// Mitsubishi GX Works2 project: ZhaoQing_OCV__5.13   PLC: Q10UDEH

TYPE ConveyorIO : STRUCT
  xUnloadCCW : BOOL;  (* 下料为反转 *)
  xUnloadAlarm : BOOL;  (* 下料报警 *)
  xUnload : BOOL;  (* 下料请求 *)
  xPutInto : BOOL;  (* 线体直接投入物料 *)
  xNotArriveAlarm : BOOL;  (* 未到达报警 *)
  xNextRun : BOOL;  (* 下段线体运行 *)
  xMotorCW : BOOL;  (* 电机正转 *)
  xMotorCCW : BOOL;  (* 电机反转 *)
  xManual : BOOL;  (* 手动 *)
  xloadCCW : BOOL;  (* 上料为反转 *)
  xLimitAlarrm : BOOL;  (* 限位报警 *)
  xLoad : BOOL;  (* 上料请求 *)
  xForward : BOOL;  (* 正转手动 *)
  xEmpty : BOOL;  (* 线体状态为空 *)
  xCWPresent : BOOL;  (* 正转检测有无传感器 *)
  xCCWPresent : BOOL;  (* 反转检测有无传感器 *)
  xBusy : BOOL;  (* 工作中 *)
  xBackward : BOOL;  (* 反转手动 *)
  xAuto : BOOL;  (* 自动 *)
  xPosLimit : BOOL;  (* 正限位 *)
  xNegLimit : BOOL;  (* 负限位 *)
  xOverWidthAlarm : BOOL;  (* 超宽报警 *)
  xError : BOOL;  (* 报警 *)
  iProductCategoryIn : INT;  (* 产品类型输入 *)
  iProductCategory : INT;  (* 产品类型记录 *)
  iProductCategoryOut : INT;  (* 产品类型输出 *)
  iDeviceID : INT;  (* 设备编号 *)
  tUnloadAlarmDelay : TIME;  (* 下料报警时间设置 *)
  tLoadDelay : TIME;  (* 上料延时设置 *)
  xSizeDeficientDetect : BOOL;  (* 尺寸缺陷检测 *)
  uiTaskIDIn : WORD;  (* 任务ID输入 *)
  uiTaskID : WORD;  (* 任务ID记录 *)
  uiTaskIDOut : WORD;  (* 任务ID输出 *)
  uiDestinationAdrIn : WORD;  (* 目标地址输入 *)
  uiDestinationAdr : WORD;  (* 目标地址记录 *)
  uiDestinationAdrOut : WORD;  (* 目标地址输出 *)
END_STRUCT END_TYPE

TYPE ShuttleCarIO : STRUCT
  xReady : BOOL;  (* 准备就绪 *)
  xForward : BOOL;  (* 正转 *)
  xBackward : BOOL;  (* 反转 *)
  iCurrentPos : INT;  (* 当前位置 *)
  iDestinationPos : INT;  (* 目标位置 *)
  xCW : BOOL;  (* 正转输出 *)
  xCCW : BOOL;  (* 反转输出 *)
  xBrake : BOOL;  (* 刹车 *)
  xHomeSwitch : BOOL;  (* 零位接近开关 *)
  xPosLimit : BOOL;  (* 正限位 *)
  xNegLimit : BOOL;  (* 负限位 *)
  xMDIExe : BOOL;  (* MDI开始 *)
  xMDIDone : BOOL;  (* MDI 完成 *)
  xPassLimit : BOOL;  (* 限位屏蔽 *)
  xPosLimitCatch : BOOL;  (* 正限位捕捉 *)
  xNegLimitCatch : BOOL;  (* 负限位捕捉 *)
  xHomeExe : BOOL;  (* 开始寻零 *)
  xHomeDone : BOOL;  (* 寻零完成 *)
  xHomeBusy : BOOL;  (* 寻零中 *)
  xHomeFailed : BOOL;  (* 寻零失败 *)
  xBusy : BOOL;  (* 工作中 *)
  tArriveDelay : TIME;  (* 到位延时 *)
  xCylinder : BOOL;  (* 气缸控制 *)
  tBrakeDelay : TIME;  (* 抱闸延时 *)
  xPauseRamp : BOOL;  (* 暂停减速斜坡标志位 *)
  xPresentDetect1 : BOOL;  (* 物料有无检测1 *)
  xPresentDetect2 : BOOL;  (* 物料有无检测2 *)
  xOvertimeAlarm : BOOL;  (* 超时报警 *)
  tSetOverTime : TIME;  (* 设置超时时间 *)
  xLooseDetect : BOOL;  (* 松绳检测 *)
  xLooseAlarm : BOOL;  (* 松绳报警 *)
END_STRUCT END_TYPE

TYPE SwitchIO : STRUCT
  xLiftCylinderRetractDetect : BOOL;
  xLiftCylinderExtendDetect : BOOL;
  xLiftCylinderRetract : BOOL;
  xLiftCylinderExtend : BOOL;
  xEntryBarCylinderRetract : BOOL;
  xLiftCylinderExtendInit : BOOL;
  xEntryEnable : BOOL;
  xExitEnable : BOOL;
  xExitBarCylinderRetract : BOOL;
  xSwithEnable : BOOL;
  xLiftCylinderRetractButton : BOOL;
  xLiftCylinderExtendButton : BOOL;
  xEntryBarCylinderRetractButton : BOOL;
  xExitBarCylinderRetractButton : BOOL;
  xPutInto : BOOL;  (* 单体复位 *)
  tSetOvertime : TIME;  (* 设定超时报警时间 *)
  xOvertimeAlarm : BOOL;  (* 超时报警 *)
END_STRUCT END_TYPE

TYPE BarCylinderIO : STRUCT
  xBarCylinderButton : BOOL;  (* 阻挡气缸 *)
  xPresentSwitch : BOOL;  (* 行程开关 *)
  xBarCylinder : BOOL;  (* 阻挡气缸 *)
  xLoad : BOOL;  (* 上料 *)
  xEmpty : BOOL;  (* 为空指示 *)
  xNextRun : BOOL;  (* 下位设备开始运行 *)
  xUnload : BOOL;  (* 下料 *)
  xTransportMotorCWButton : BOOL;  (* 输送电机正转按钮 *)
  xTransportMotorCW : BOOL;  (* 输送电机正转 *)
  xTransportMotorCCWButton : BOOL;  (* 输送电机反转按钮 *)
  xTransportMotorCCW : BOOL;  (* 输送电机反转 *)
  iProductCategory : INT;  (* 产品种类 *)
  tLoadDelay : TIME;  (* 上料延时 *)
END_STRUCT END_TYPE

// global labels: Global1
VAR_GLOBAL
  g_xAuto AT M11 : BOOL;
  g_xManual : BOOL;
  g_xEStop AT X0BC : BOOL;
  g_xReset AT X0BE : BOOL;
  g_xStackLampRed AT Y2C1 : BOOL;
  g_xStackLampAmber AT Y2C3 : BOOL;
  g_xStackLampGreen AT Y2C2 : BOOL;
  g_xBuzzer AT Y2C4 : BOOL;
  g_xStop AT M2 : BOOL;
  g_xLocalAutoStart AT M1 : BOOL;
  g_xRemoteAutoStart AT M0 : BOOL;
  g_xRemoteAuto AT M10 : BOOL;
  g_iState AT D40 : INT;
  g_iLocalAutoStep : BOOL;
  g_xAlarm : BOOL;
  g_xPause AT M3 : BOOL;  (* 暂停 *)
  g_iDeviceIDSelect AT D0 : INT;
  g_xImport1Force AT M165 : BOOL;
  g_xImport2Force AT M166 : BOOL;
  g_xImport3Force AT M167 : BOOL;
  g_xResetSingle AT M4 : BOOL;  (* 单线体复位 *)
  g_xInsertTask AT M5 : BOOL;  (* 插入任务 *)
  g_iInsertTask AT D2 : INT;  (* 插入任务号 *)
  g_iConveyorStatus AT D4 : INT;
  g_xChenPinComFailed AT M168 : BOOL;
END_VAR

// task Task_01 (event TRUE, interval 0, priority 31): POU, Start, tcp

FUNCTION_BLOCK Conveyor
VAR
  m_xPresentDelay : BOOL;  (* 有无判断延时 *)
  m_xLoadDelayOut : BOOL;  (* 上料延时输出 *)
  m_xInitial : BOOL;  (* 初始化 *)
  m_tUnloadTimer : TIME;  (* 下料计时器 *)
  m_tPresentDelayCurrentTime : TIME;
  m_tonUnloadAlam : TON;  (* 下料报警定时器 *)
  m_tonPresentDelay : TON;  (* 物料有无判断延时，防止误动作 *)
  m_tonNotArriveAlarm : TON;  (* 未到达报警计时 *)
  m_tonLoadDelay : TON;  (* 上料延时 *)
  m_tNotArriveCurrentTime : TIME;  (* 未到达报警计时当前时间 *)
  m_tLoadTimer : TIME;  (* 上料计时器 *)
  iStep : INT;  (* 上料步骤 *)
  m_wStateWord : INT;
END_VAR
VAR_IN_OUT
  ConveyorMotor : ConveyorIO;  (* 输送线输入输出 *)
END_VAR
(*////////////////////////////////////////////////////////////////////////////////////////////////////////////
//传输线控制FB块，可控制单方向线体，双向旋转线体，支持双向上下料            
//线体初始化后为空的情况下输入xLoad信号即可进行上料动作，使用xLoadCCW信号可反方向上料
//增加了产品信息和产品种类的储存，当传输线为空和上料进行标志位为零的情况下清除产品信息和产品种类
//使用方式是在置位xLoad信号后，把产品信息和产品种类传入，等下料后自动清零
//线体不为空的情况下使用xUnload信号可进行下料动作，物料有无传感器的下降沿后出发计时器，延时断开传输线旋转
//单方向传输线体把xLoadCCW、xUnloadCCW设置为零，双向线体上料方向和下料反向的,方向固定的 把xUnloadCCW设置为1
//双方向线体双向都能上下料的要根据上料的方向来设置xLoadCCW,xUnloadCCW
//增加工作中信号xBusy当电机正转 显示为工作中
//增加上下料超时报警，xLoadAlarm，xUnloadAlarm，设定时间在LOAD_UNLOAD_TIME常量上，现在设置的为30秒
//增加xPutInto信号，用于直接投入的物料，检测开关感应到后，直接进入下料流程，上升沿有效
//离开延时改为变量 iLeaveDelay 默认为0 离开检测开关离输送线尾端比较远的线体需要根据情况设定100ms为单位
//增加初始化标志位，增加进入延时时间，初始化为进入延时时间为0 ，离开延时时间为2S，通过外围接口可以更改
//修改信息  修改后请增加版本
//12-17进行了优化，增加了未到达报警，当物料未传送到下一设备，就报未到达报警，使用xNextRun标志位制作，没有正常到达
//第0步，不能跳转到第一步把标志位复位，即出现中断情况，2秒后报警
//修改信息  修改后请增加版本
上料延时增加为50ms防止干扰信号
nextrun信号在 第三步也要复位
增加限位报警
增加超宽报警
增加产品型号输出在下料的时候把产品型号输送给下一段线体
增加线体单独复位
增加任务插入功能配合全局变量
增加暂停功能
增加线体状态字显示  0 空闲 1：有料  2 工作中  3  超限报警 4 超宽报警  5 未到达报警  6 下料超时报警
空料判断放在自动前，进行有无报警判断，然后跳转
//YAO      V1.0
///////////////////////////////////////////////////////////////////////////////////////////////////////////
(*********************************************************)
(*//初始化，
//上料延时位0S，下料报警延时为30S
//下料延时设一个比较大的时间，主要依靠xunload标志位来停止输送线，特殊情况可以用延时来停止物流线下料
//设置时间大的时候计时器会失效*)
IF NOT m_xInitial THEN
	ConveyorMotor.tLoadDelay:=T#100ms;
	ConveyorMotor.tUnloadAlarmDelay:=T#30s;
	ConveyorMotor.xPosLimit:=1;
	ConveyorMotor.xNegLimit:=1;
	ConveyorMotor.xSizeDeficientDetect:=0;
	m_xInitial:=1;
END_IF;
(*//自动
//复位信号把步号置0，但xLoad与xUnload没有复位，调用程序需要注意复位后把这两个信号置零，以免发生误动作
//物料有无判断增加延时，防止开自动瞬间误动作发生*)
m_tonPresentDelay(IN:= ConveyorMotor.xCWPresent OR ConveyorMotor.xCCWPresent,
                  PT:=T#100ms,
				  Q:= m_xPresentDelay,
				  ET:= m_tPresentDelayCurrentTime);
CASE iStep OF
	0:(*//初始化*)
	ConveyorMotor.xMotorCW:=0;
	ConveyorMotor.xMotorCCW:=0;
	ConveyorMotor.iProductCategoryOut:=0;
	ConveyorMotor.uiTaskIDOut:=0;
	ConveyorMotor.uiDestinationAdOut:=0;
(*	//判断物料有无传感器*)	
		IF m_xPresentDelay THEN			
			ConveyorMotor.xEmpty:=0;
			IF g_xAuto AND NOT ConveyorMotor.xError THEN(*//自动情况下进行跳转*)(*无超限报警*)
				iStep:=3;
			END_IF;
		ELSE
			ConveyorMotor.xEmpty:=1;
			IF g_xAuto AND NOT ConveyorMotor.xError THEN(*//自动情况下进行跳转*)(*无超限报警*)
				iStep:=1;	
			END_IF;		
	END_IF;	
	1: (*//上料*)
	ConveyorMotor.xNextRun:=0;
	IF ConveyorMotor.xLoad    THEN (*//上料开始*)
		ConveyorMotor.iProductCategory:=0;	(*//上料开始清除产品信息*)
		ConveyorMotor.uiTaskID:=0;
		ConveyorMotor.uiDestinationAdr:=0;		
		iStep:=2;		
	END_IF;
	2: (*//上料完成*)
	ConveyorMotor.iProductCategory:=ConveyorMotor.iProductCategoryIn;(* //产品信息传入*)		
	ConveyorMotor.uiTaskID:=ConveyorMotor.uiTaskIDIn;
	ConveyorMotor.uiDestinationAdr:=ConveyorMotor.uiDestinationAdrIn;
	IF ConveyorMotor.xloadCCW THEN
		ConveyorMotor.xMotorCCW:=1; 
		ConveyorMotor.xMotorCW:=0;
	ELSE
	    ConveyorMotor.xMotorCW:=1;  
		ConveyorMotor.xMotorCCW:=0;
	END_IF;
		m_tonLoadDelay(IN:= (ConveyorMotor.xCWPresent AND NOT ConveyorMotor.xloadCCW) 
		                                        OR (ConveyorMotor.xCCWPresent AND ConveyorMotor.xloadCCW) ,
		                               PT:= ConveyorMotor.tLoadDelay ,
		                               Q:= m_xLoadDelayOut ,
		                               ET:= m_tLoadTimer );
	    IF (m_xLoadDelayOut AND NOT ConveyorMotor.xSizeDeficientDetect)   (*无尺寸检测时  只检测一个开关*)
	    	OR (m_xLoadDelayOut AND ConveyorMotor.xSizeDeficientDetect(*有尺寸检测时  要检测两个开关*)
	    	                                          AND ConveyorMotor.xCCWPresent 
	    	                                          AND ConveyorMotor.xCWPresent)      THEN 	 
		    iStep:=3;
			    ELSIF (m_xLoadDelayOut 
		                       AND ConveyorMotor.xSizeDeficientDetect(*尺寸不足报警*)
	    	                  AND (NOT ConveyorMotor.xCCWPresent OR NOT ConveyorMotor.xCWPresent))  
	    THEN
	    	    ConveyorMotor.xOverWidthAlarm:=1;
	    	   iStep:=0;               
	    END_IF;

	3:(*//下料请求*)	
	ConveyorMotor.xMotorCW:=0;
	ConveyorMotor.xMotorCCW:=0;
	ConveyorMotor.xEmpty:=0;
	IF ConveyorMotor.xUnload AND NOT ConveyorMotor.xOverWidthAlarm  THEN (*无超宽报警可以下料*)
		iStep:=4;
	END_IF;
	4:(*	//下料完成*)
	IF ConveyorMotor.xUnloadCCW THEN   
		ConveyorMotor.xMotorCCW:=1;  
		ConveyorMotor.xMotorCW:=0;
		ELSE
	    ConveyorMotor.xMotorCW:=1;  
		ConveyorMotor.xMotorCCW:=0;
	END_IF;
	ConveyorMotor.xNextRun:=1; (*下一段线体旋转*)
	ConveyorMotor.iProductCategoryOut:=ConveyorMotor.iProductCategory;(*产品型号输出给下一段线体*)
	ConveyorMotor.uiDestinationAdrOut:=ConveyorMotor.uiDestinationAdr;
	ConveyorMotor.uiTaskIDOut:=
	IF NOT ConveyorMotor.xUnload THEN 
		istep:=0;
	END_IF;
END_CASE;
(*投入上料，搬出下料，也可用来初始化*)
IF LDP(TRUE,ConveyorMotor.xPutInto) THEN
	iStep:=0;
END_IF;
(*//当前任务显示*)
IF LDP(TRUE,ConveyorMotor.iDeviceID=g_iDeviceIDSelect) THEN
	g_iInsertTask:=ConveyorMotor.iProductCategory;
END_IF;
	(*//插入任务*)
IF g_xInsertTask AND ConveyorMotor.iDeviceID=g_iDeviceIDSelect THEN
	ConveyorMotor.iProductCategory:=g_iInsertTask;
END_IF;
(*//单线体复位，当设备号与本线体一致的时候执行复位*)
IF (g_xResetSingle AND ConveyorMotor.iDeviceID=g_iDeviceIDSelect)THEN (* //非正常情况下切断xNextRun不会复位，通过这个标志位会出发报警*)(*增加单体复位*)
	iStep:=0;
	ConveyorMotor.xNextRun:=0; 
	ConveyorMotor.xLimitAlarrm:=0;
	ConveyorMotor.xOverWidthAlarm:=0;
END_IF;
(*//手动*)
IF g_xManual THEN
(*	iStep:=0; *)(*//手动后上下料程序步骤清零*)
	(*//正转*)
	IF ConveyorMotor.xForward 
		AND ConveyorMotor.xBackward=0 
		AND ConveyorMotor.xMotorCCW=0 
		AND g_xEStop THEN
		ConveyorMotor.xMotorCW:=1;
		ConveyorMotor.xMotorCCW:=0;
		ELSE
		ConveyorMotor.xMotorCW:=0;
	END_IF;
	(*//反转*)
	IF ConveyorMotor.xBackward 
		AND ConveyorMotor.xForward=0 
		AND ConveyorMotor.xMotorCW=0 
		AND g_xEStop THEN
		ConveyorMotor.xMotorCCW:=1;
		conveyormotor.xMotorCW:=0;
		ELSE
		ConveyorMotor.xMotorCCW:=0;
	END_IF;
END_IF;
(*暂停*)
IF g_xPause THEN
	ConveyorMotor.xMotorCCW:=0;
	ConveyorMotor.xMotorCW:=0;
END_IF;
(*工作中信号输出*)
ConveyorMotor.xBusy:=ConveyorMotor.xMotorCCW OR ConveyorMotor.xMotorCW;
(*//未到达报警*)
m_tonNotArriveAlarm(IN:= iStep=0 AND ConveyorMotor.xNextRun  ,PT:= T#2s,Q:= ConveyorMotor.xNotArriveAlarm ,ET:= m_tNotArriveCurrentTime );
(*//下料超时报警*)
m_tonUnloadAlam(IN:= iStep=4,PT:=ConveyorMotor.tUnloadAlarmDelay,Q:= ConveyorMotor.xUnloadAlarm,ET:=m_tUnloadTimer );
(*//限位报警,进料检测开关失效*)
IF ( ((ConveyorMotor.xloadCCW AND NOT ConveyorMotor.xNegLimit)            (*反转上料，碰到负限位*)
	OR  ( NOT ConveyorMotor.xloadCCW AND NOT ConveyorMotor.xPosLimit)) (*正转上料，碰到正限位*)
    AND iStep=2) (*上料过程*)
    OR
   ( iStep=4 (*下料过程*)
	AND( (ConveyorMotor.xUnloadCCW AND NOT ConveyorMotor.xPosLimit)  
	OR (NOT ConveyorMotor.xUnloadCCW AND NOT ConveyorMotor.xNegLimit)))    
    THEN
    ConveyorMotor.xLimitAlarrm:=1;
    iStep:=0;
END_IF;
(*//超宽报警*)
IF iStep=3 AND (NOT ConveyorMotor.xNegLimit OR NOT ConveyorMotor.xPosLimit) THEN
	ConveyorMotor.xOverWidthAlarm:=1;
END_IF;
(*//总报警*)
ConveyorMotor.xError:=ConveyorMotor.xLimitAlarrm
                                              OR ConveyorMotor.xNotArriveAlarm
                                              OR ConveyorMotor.xUnloadAlarm                                             
                                              OR ConveyorMotor.xOverWidthAlarm;

(*//状态输出*)(*状态显示，容易造成指针容量不足*)
IF ConveyorMotor.xEmpty AND NOT ConveyorMotor.xBusy THEN
	m_wStateWord:=0;
END_IF;
IF ConveyorMotor.xEmpty=0 THEN
		m_wStateWord:=1;
END_IF;
IF ConveyorMotor.xBusy THEN
		m_wStateWord:=2;
END_IF;
IF ConveyorMotor.xLimitAlarrm THEN
		m_wStateWord:=3;
END_IF;
IF ConveyorMotor.xOverWidthAlarm THEN
		m_wStateWord:=4;
END_IF;
(*IF ConveyorMotor.xNotArriveAlarm THEN	
		m_wStateWord:=5;
END_IF;*)
IF ConveyorMotor.xUnloadAlarm THEN
		m_wStateWord:=6;	
END_IF;
(*选择本线体后，将状态赋值给全局变量进行显示*)
IF ConveyorMotor.iDeviceID=g_iDeviceIDSelect THEN
	g_iConveyorStatus:=m_wStateWord;
END_IF;
END_FUNCTION_BLOCK

PROGRAM POU
VAR
  Cylinder12309 : ShuttleCar;
  CylinderIO12309 : ShuttleCarIO;
  ConveyorIO12114 : ConveyorIO;
  Conveyor12114 : Conveyor;
  Conveyor12115 : Conveyor;
  ConveyorIO12115 : ConveyorIO;
  Switch12312 : Switch;
  SwitchIO12312 : SwitchIO;
  Conveyor12123 : Conveyor;
  ConveyorIO12123 : ConveyorIO;
  Conveyor12124 : Conveyor;
  ConveyorIO12124 : ConveyorIO;
  Conveyor12125 : Conveyor;
  ConveyorIO12125 : ConveyorIO;
  Switch12203 : Switch;
  SwitchIO12203 : SwitchIO;
  Conveyor12142 : Conveyor;
  ConveyorIO12142 : ConveyorIO;
  Bar12326 : BarCylinder;
  BarIO12326 : BarCylinderIO;
  Conveyor12116 : Conveyor;
  ConveyorIO12116 : ConveyorIO;
  Cylinder12308 : ShuttleCar;
  CylinderIO12308 : ShuttleCarIO;
  Conveyor12111 : Conveyor;
  ConveyorIO12111 : ConveyorIO;
  Conveyor12112 : Conveyor;
  ConveyorIO12112 : ConveyorIO;
  Switch12311 : Switch;
  SwitchIO12311 : SwitchIO;
  Conveyor12113 : Conveyor;
  ConveyorIO12113 : ConveyorIO;
  Conveyor12120 : Conveyor;
  ConveyorIO12120 : ConveyorIO;
  Conveyor12121 : Conveyor;
  ConveyorIO12121 : ConveyorIO;
  Conveyor12122 : Conveyor;
  ConveyorIO12122 : ConveyorIO;
  Cylinder12307 : ShuttleCar;
  CylinderIO12307 : ShuttleCarIO;
  Conveyor12108 : Conveyor;
  ConveyorIO12108 : ConveyorIO;
  Conveyor12109 : Conveyor;
  ConveyorIO12109 : ConveyorIO;
  Switch12310 : Switch;
  SwitchIO12310 : SwitchIO;
  Conveyor12110 : Conveyor;
  ConveyorIO12110 : ConveyorIO;
  Conveyor12117 : Conveyor;
  ConveyorIO12117 : ConveyorIO;
  Conveyor12118 : Conveyor;
  ConveyorIO12118 : ConveyorIO;
  Conveyor12119 : Conveyor;
  ConveyorIO12119 : ConveyorIO;
  Conveyor12203 : Conveyor;
  ConveyorIO12203 : ConveyorIO;
  Conveyor12143 : Conveyor;
  ConveyorIO12143 : ConveyorIO;
  Switch12330 : Switch;
  ConveyorIO12144 : ConveyorIO;
  ConveyorIO12333 : ConveyorIO;  (* OCV2顶升移载进入线体 *)
  ConveyorIO12152 : ConveyorIO;  (* OCV2顶升移载离开线体 *)
  SwitchIO12333 : SwitchIO;  (* OCV2顶升移载 *)
  m_xTS1ExportPermit : BOOL;  (* OCV2顶升移载 *)
  m_xConveyor12114Export : BOOL;  (* 12114线体输出 *)
  ConveyorIO12146 : ConveyorIO;
  m_xTS2ExportPermit : BOOL;
  m_xMotorFlag : BOOL;
  m_xTS3ExportPermit : BOOL;
  SwitchIO12330 : SwitchIO;
  Switch12333 : Switch;  (* OCV2顶升移载 *)
  SwitchIO12321 : SwitchIO;
  Switch12321 : Switch;  (* OCV2顶升移载 *)
  Conveyor12141 : Conveyor;
  ConveyorIO12141 : ConveyorIO;
  Conveyor12140 : Conveyor;
  ConveyorIO12140 : ConveyorIO;
  m_iSwitch12321Select : INT;
  Conveyor12138 : Conveyor;
  ConveyorIO12138 : ConveyorIO;
  Conveyor12139 : Conveyor;
  ConveyorIO12139 : ConveyorIO;
  Conveyor12136 : Conveyor;
  ConveyorIO12136 : ConveyorIO;
  Conveyor12137 : Conveyor;
  ConveyorIO12137 : ConveyorIO;
  Switch12317 : Switch;
  SwitchIO12317 : SwitchIO;
  ConveyorIO12135 : ConveyorIO;
  ConveyorIO12134 : ConveyorIO;
  m_iSwitch12317Select : INT;
  Conveyor12132 : Conveyor;
  ConveyorIO12132 : ConveyorIO;
  Conveyor12133 : Conveyor;
  ConveyorIO12133 : ConveyorIO;
  Conveyor12131 : Conveyor;
  ConveyorIO12131 : ConveyorIO;
  Conveyor12130 : Conveyor;
  ConveyorIO12130 : ConveyorIO;
  Switch12314 : Switch;
  SwitchIO12314 : SwitchIO;
  Conveyor12129 : Conveyor;
  ConveyorIO12129 : ConveyorIO;
  Conveyor12128 : Conveyor;
  ConveyorIO12128 : ConveyorIO;
  m_iSwitch12314Select : INT;
  Conveyor12126 : Conveyor;
  ConveyorIO12126 : ConveyorIO;
  Conveyor12127 : Conveyor;
  ConveyorIO12127 : ConveyorIO;
  Cylinder12320 : ShuttleCar;
  CylinderIO12320 : ShuttleCarIO;
  Cylinder12316 : ShuttleCar;
  CylinderIO12316 : ShuttleCarIO;
  Cylinder12313 : ShuttleCar;
  CylinderIO12313 : ShuttleCarIO;
  Conveyor12147 : Conveyor;
  ConveyorIO12147 : ConveyorIO;
  Conveyor12148 : Conveyor;
  ConveyorIO12148 : ConveyorIO;
  Lifter8 : ShuttleCar;
  Lifter8IO : ShuttleCarIO;
  Lifter8Speed : ShuttleCarVelocityFB;
  Conveyor8 : Conveyor;
  Conveyor8IO : ConveyorIO;
  Lifter9 : ShuttleCar;
  Lifter9IO : ShuttleCarIO;
  Lifter9Speed : ShuttleCarVelocityFB;
  Conveyor9 : Conveyor;
  Conveyor9IO : ConveyorIO;
  Conveyor12156 : Conveyor;
  ConveyorIO12156 : ConveyorIO;
  Conveyor12155 : Conveyor;
  ConveyorIO12155 : ConveyorIO;
  m_tonSwitch1NOSeleteDelay : TON;
  m_tonSwitch2NOSeleteDelay : TON;
  m_tonSwitch3NOSeleteDelay : TON;
  m_xSwitch12321NoSeleteDelay : BOOL;
  m_xSwitch12317NoSeleteDelay : BOOL;
  m_xSwitch12314NoSeleteDelay : BOOL;
  m_tSwitch12321NOSeleteCurrent : TIME;
  m_tSwitch12317NOSeleteCurrent : TIME;
  m_tSwitch12314NOSeleteCurrent : TIME;
  Switch12312Priority : PriorityFB;
  m_xSwitch12312Task : INT;
  Conveyor12159 : Conveyor;
  ConveyorIO12159 : ConveyorIO;
  Switch12337 : Switch;
  SwitchIO12337 : SwitchIO;
  ConveyorIO12158 : ConveyorIO;
  ConveyorIO12157 : ConveyorIO;
  ConveyorIO12321 : ConveyorIO;
  Switch12311Priority : PriorityFB;
  m_xSwitch12311Task : INT;
  SwitchIO12204 : SwitchIO;
  Switch12204 : Switch;
  ConveyorIO12145 : ConveyorIO;
  ConveyorIO12204 : ConveyorIO;
  Conveyor12151 : Conveyor;
  ConveyorIO12151 : ConveyorIO;
  Conveyor12150 : Conveyor;
  ConveyorIO12150 : ConveyorIO;
  Conveyor12149 : Conveyor;
  ConveyorIO12149 : ConveyorIO;
  Switch12328 : Switch;
  SwitchIO12328 : SwitchIO;
  Lifter8Priority : PriorityFB;
  m_iLifter8Task : INT;
  m_xSwitch12321Select : BOOL;
  m_xSwitch12317Select : BOOL;
  Cylinder12301 : ShuttleCar;
  CylinderIO12301 : ShuttleCarIO;
  Cylinder12302 : ShuttleCar;
  CylinderIO12302 : ShuttleCarIO;
  Cylinder12303 : ShuttleCar;
  CylinderIO12303 : ShuttleCarIO;
  Cylinder12304 : ShuttleCar;
  CylinderIO12304 : ShuttleCarIO;
  Conveyor12101 : Conveyor;
  ConveyorIO12101 : ConveyorIO;
  Conveyor12102 : Conveyor;
  ConveyorIO12102 : ConveyorIO;
  Conveyor12103 : Conveyor;
  ConveyorIO12103 : ConveyorIO;
  Conveyor12104 : Conveyor;
  ConveyorIO12104 : ConveyorIO;
  ShuttleCar12401 : ShuttleCar;
  ShuttleCarIO12401 : ShuttleCarIO;
  Conveyor12105 : Conveyor;
  ConveyorIO12105 : ConveyorIO;
  Conveyor12106 : Conveyor;
  ConveyorIO12106 : ConveyorIO;
  Switch12201 : Switch;
  SwitchIO12201 : SwitchIO;
  Switch12202 : Switch;
  SwitchIO12202 : SwitchIO;
  Conveyor12201 : Conveyor;
  ConveyorIO12201 : ConveyorIO;
  Conveyor12202 : Conveyor;
  ConveyorIO12202 : ConveyorIO;
  Conveyor12401 : Conveyor;
  ConveyorIO12401 : ConveyorIO;
  Rotor12501 : ShuttleCar;
  RotorIO12501 : ShuttleCarIO;
  Conveyor12501 : Conveyor;
  ConveyorIO12501 : ConveyorIO;
  Conveyor12154 : Conveyor;
  ConveyorIO12154 : ConveyorIO;
  ShuttleCar12401Position : ARRAY [0..5] OF INT;
  ii : INT;
  ConveyorIO12107 : ConveyorIO;
  m_xSwitch12314Select : BOOL;
  Conveyor12146 : Conveyor;
  Switch12330ConveyorOut : ConveyorIO;
  m_xPickOutDone : BOOL;  (* 分拣完成 *)
  ConveyorIO12160 : ConveyorIO;  (* OCV1工位 *)
  m_xOCV1Done : BOOL;  (* OCV1完成 *)
  Conveyor12160 : Conveyor;
  Conveyor12161 : Conveyor;
  ConveyorIO12161 : ConveyorIO;
  ConveyorIO12162 : ConveyorIO;
  Conveyor12162 : Conveyor;
  TonScan1 : TON;
  TonScan1Time : TIME;
  TonScan2 : TON;
  TonScan2Time : TIME;
  xTonScan1 : BOOL;
  xTonScan2 : BOOL;
END_VAR
IF M1 AND M2 THEN D333:=D333;END_IF;
(*提升机8*)
Lifter8(ShuttleCarInOut:=Lifter8IO);
(*ShuttleCarCurrentPosition(XC2 OR XC4 OR XC3 ,XC2 ,XC3, XC4, Lifter8IO.iCurrentPos);*)
IF XC1 AND XC2 THEN
	Lifter8IO.iCurrentPos:=1;
ELSIF XC2 AND NOT XC1 THEN
	Lifter8IO.iCurrentPos:=2;
ELSIF XC3 THEN
	Lifter8IO.iCurrentPos:=3;
ELSIF XC4 THEN
	Lifter8IO.iCurrentPos:=4;
END_IF;
Lifter8Speed(xEnable:= g_xAuto,
                        xMotorCW:= Lifter8IO.xCW ,
                        xMotorCCW:= Lifter8IO.xCCW,
                        xPosition1Switch:= XC2 OR XC4,
                        xDecelerationSwitch:= XC0 ,
	                    xPosition2Switch:= XC3 ,
	                   xHighSpeed:= Y296 );
Lifter8IO.xReady:=XBA;
Lifter8IO.xLooseDetect:=XC6;;
Lifter8IO.xForward:=M107 OR XC7;
Lifter8IO.xBackward:=M108 OR XC8;
Lifter8IO.xPosLimit:=XBF;
Lifter8IO.xNegLimit:=XC5;
Y294:=Lifter8IO.xCW;
Y295:=Lifter8IO.xCCW;
Y299:=Lifter8IO.xBrake;
Lifter8IO.tArriveDelay:=T#500ms;

Conveyor8(ConveyorMotor:=Conveyor8IO);
Conveyor8IO.xForward:=M109;
Conveyor8IO.xBackward:=M110;
Conveyor8IO.xCWPresent:=XC9;
Conveyor8IO.xCCWPresent:=XCA;
Y29A:=Conveyor8IO.xMotorCW;
Y29B:=Conveyor8IO.xMotorCCW;
Conveyor8IO.xSizeDeficientDetect:=1;
Conveyor8IO.iDeviceID:=8;

(*提升机9*)
Lifter9(ShuttleCarInOut:=Lifter9IO);
ShuttleCarCurrentPosition(XCC OR XCD ,XCC ,XCD,FALSE, Lifter9IO.iCurrentPos);
Lifter9Speed(xEnable:= g_xAuto,
                        xMotorCW:= Lifter9IO.xCW ,
                        xMotorCCW:=Lifter9IO.xCCW,
                        xPosition1Switch:= XCC,
                        xDecelerationSwitch:= XCB,
	                    xPosition2Switch:= XCD ,
	                    xHighSpeed:= Y2A1 );
Lifter9IO.xReady:=XBB;
Lifter9IO.xForward:=M111 OR XD1;
Lifter9IO.xBackward:=M112 OR XD2;
Lifter9IO.xLooseDetect:=XD0;
Lifter9IO.xPosLimit:=XCE;
Lifter9IO.xNegLimit:=XCF;
Y29F:=Lifter9IO.xCW;
Y2A0:=Lifter9IO.xCCW;
Y2A4:=Lifter9IO.xBrake;

Conveyor9(ConveyorMotor:=Conveyor9IO);
Conveyor9IO.xForward:=M113;
Conveyor9IO.xBackward:=M114;
Conveyor9IO.xCWPresent:=XD4;
Conveyor9IO.xCCWPresent:=XD3;
Y2A6:=Conveyor9IO.xMotorCW;
Y2A5:=Conveyor9IO.xMotorCCW;
Conveyor9IO.iDeviceID:=9;
(*H750高温库人工换内衬线体*)
(*高位库2巷道入库*)
Cylinder12301(ShuttleCarInOut:=CylinderIO12301);
ShuttleCarCurrentPosition( X3 OR X4 ,X4 ,X3, FALSE, CylinderIO12301.iCurrentPos );
CylinderIO12301.xForward:=M137;
CylinderIO12301.xBackward:=M138;
CylinderIO12301.xCylinder:=1;
Y201:=CylinderIO12301.xCW;
Y202:=CylinderIO12301.xCCW;
CylinderIO12301.xPresentDetect1:=X02;

Conveyor12101(ConveyorMotor:=ConveyorIO12101);
ConveyorIO12101.xForward:=M139;
ConveyorIO12101.xCWPresent:=X1;
Y203:=ConveyorIO12101.xMotorCW;
M362:= NOT ConveyorIO12101.xEmpty;
M363:=ConveyorIO12101.xError;
ConveyorIO12101.iDeviceID:=12101;

(*高位库2巷道出库*)
Cylinder12302(ShuttleCarInOut:=CylinderIO12302);
ShuttleCarCurrentPosition( X6 OR X7 ,X7,X6, FALSE, CylinderIO12302.iCurrentPos );
CylinderIO12302.xForward:=M140;
CylinderIO12302.xBackward:=M141;
CylinderIO12302.xCylinder:=1;
Y204:=CylinderIO12302.xCW;
Y205:=CylinderIO12302.xCCW;
CylinderIO12302.xPresentDetect1:=X05;

Conveyor12102(ConveyorMotor:=ConveyorIO12102);
ConveyorIO12102.xForward:=M141;
ConveyorIO12102.xCWPresent:=X8;
Y206:=ConveyorIO12102.xMotorCW;
M410:= NOT conveyorIO12102.xEmpty;
M411:= ConveyorIO12102.xError;
ConveyorIO12102.iDeviceID:=12102;

(*高位库1巷道出库*)
Cylinder12303(ShuttleCarInOut:=CylinderIO12303);
ShuttleCarCurrentPosition( X9 OR XA ,XA,X9, FALSE, CylinderIO12303.iCurrentPos );
CylinderIO12303.xForward:=M142;
CylinderIO12303.xBackward:=M143;
CylinderIO12303.xCylinder:=1;
Y207:=CylinderIO12303.xCW;
Y208:=CylinderIO12303.xCCW;
CylinderIO12303.xPresentDetect1:=X0B;

Conveyor12103(ConveyorMotor:=ConveyorIO12103);
ConveyorIO12103.xForward:=M144;
ConveyorIO12103.xCWPresent:=XC;
M412:= NOT conveyorIO12103.xEmpty;
M413:= ConveyorIO12103.xError;
ConveyorIO12103.iDeviceID:=12103;
Y209:=ConveyorIO12103.xMotorCW;

(*高位库1巷道入库*)
Cylinder12304(ShuttleCarInOut:=CylinderIO12304);
ShuttleCarCurrentPosition( XF OR X10 ,X10,XF, FALSE, CylinderIO12304.iCurrentPos );
CylinderIO12304.xForward:=M145;
CylinderIO12304.xBackward:=M146;
CylinderIO12304.xCylinder:=1;
Y21A:=CylinderIO12304.xCW;
Y21B:=CylinderIO12304.xCCW;
CylinderIO12304.xPresentDetect1:=X0E;

Conveyor12104(ConveyorMotor:=ConveyorIO12104);
ConveyorIO12104.xForward:=M144;
ConveyorIO12104.xCWPresent:=XD;
Y21C:=ConveyorIO12104.xMotorCW;
M414:= NOT conveyorIO12104.xEmpty;
M415:= ConveyorIO12104.xError;
ConveyorIO12104.iDeviceID:=12104;

(*高位库RGV*)
(*ShuttleCar12401(ShuttleCarInOut:= ShuttleCarIO12401 );
ShuttleCar12401Position[0]:=1;
ShuttleCar12401Position[1]:=1;
ShuttleCar12401Position[2]:=1;
ShuttleCar12401Position[3]:=1;
ShuttleCar12401Position[4]:=1;
ShuttleCar12401Position[5]:=1;

Y2CA:=ShuttleCarVelocityEncoder( g_xAuto , D190 , ShuttleCar12401Position[ShuttleCarIO12401.iDestinationPos] );
IF LDP(TRUE,g_xAuto) THEN
	ShuttleCarIO12401.iCurrentPos:=0;
END_IF;
FOR ii:=0 TO 5 BY 1 DO
	IF abs(D190-ShuttleCar12401Position[ii])<10 THEN
		ShuttleCarIO12401.iCurrentPos:=ii;
	END_IF;
END_FOR;

ShuttleCarIO12401.xReady:=XBD;
ShuttleCarIO12401.xForward:=M147 OR XD5;
ShuttleCarIO12401.xBackward:=M148 OR XD6;
ShuttleCarIO12401.xPosLimit:=XDA;
ShuttleCarIO12401.xNegLimit:=XDB;
Y2C8:=ShuttleCarIO12401.xCW;
Y2C9:=ShuttleCarIO12401.xCCW;
Y2BD:=ShuttleCarIO12401.xBrake;

Conveyor12105(ConveyorMotor:=ConveyorIO12105);
ConveyorIO12105.xForward:=M149;
ConveyorIO12105.xCWPresent:=X11;
Y21D:=ConveyorIO12105.xMotorCW;
M416:= NOT conveyorIO12105.xEmpty;
M417:= ConveyorIO12105.xError;
ConveyorIO12105.iDeviceID:=12105;

Conveyor12106(ConveyorMotor:=ConveyorIO12106);
ConveyorIO12106.xForward:=M150;
ConveyorIO12106.xCWPresent:=X12;
Y21E:=ConveyorIO12106.xMotorCW;
M418:= NOT conveyorIO12106.xEmpty;
M419:= ConveyorIO12106.xError;
ConveyorIO12106.iDeviceID:=12106;

Switch12202(ConveyorEntryIO:=ConveyorIO12202 ,
                                                        ConveyorExitIO:=ConveyorIO12107 ,
                                                        SwitchIO:=SwitchIO12202 );
SwitchIO12202.xLiftCylinderExtendButton:=M151;
SwitchIO12202.xLiftCylinderRetractButton:=M152;
Y220:=SwitchIO12202.xLiftCylinderExtend;
Y221:=SwitchIO12202.xLiftCylinderRetract;
SwitchIO12202.xLiftCylinderExtendDetect:=X14;
SwitchIO12202.xLiftCylinderRetractDetect:=X15;
ConveyorIO12202.xForward:=M153;
ConveyorIO12202.xCWPresent:=X13;
Y21F:=ConveyorIO12202.xMotorCW;
ConveyorIO12202.tLoadDelay:=T#3s;
M420:= NOT conveyorIO12202.xEmpty;
M421:= ConveyorIO12202.xError;
ConveyorIO12202.iDeviceID:=12202;
ConveyorIO12107.xForward:=M154;
ConveyorIO12107.xCWPresent:=X13;
Y227:=ConveyorIO12107.xMotorCW;
ConveyorIO12107.iDeviceID:=12202;

Switch12201(ConveyorEntryIO:=ConveyorIO12107 ,
                                                        ConveyorExitIO:=ConveyorIO12201 ,
                                                        SwitchIO:=SwitchIO12201 );
SwitchIO12201.xLiftCylinderExtendButton:=M155;
SwitchIO12201.xLiftCylinderRetractButton:=M156;
Y220:=SwitchIO12201.xLiftCylinderExtend;
Y221:=SwitchIO12201.xLiftCylinderRetract;
SwitchIO12201.xLiftCylinderExtendDetect:=X14;
SwitchIO12201.xLiftCylinderRetractDetect:=X15;
ConveyorIO12107.tLoadDelay:=T#3s;
ConveyorIO12201.xForward:=M157;
ConveyorIO12201.xCWPresent:=X19;
Y226:=ConveyorIO12201.xMotorCW;
M422:= NOT conveyorIO12101.xEmpty;
M423:= ConveyorIO12101.xError;
ConveyorIO12101.iDeviceID:=12201;*)

(*常温库1巷道出库线体*)
Cylinder12309(ShuttleCarInOut:=CylinderIO12309);
ShuttleCarCurrentPosition( X43 OR X44 ,X44 ,X43, FALSE, CylinderIO12309.iCurrentPos );
CylinderIO12309.xForward:=M30;
CylinderIO12309.xBackward:=M31;
CylinderIO12309.xCylinder:=1;
Y23D:=CylinderIO12309.xCW;
Y23C:=CylinderIO12309.xCCW;
CylinderIO12309.xPresentDetect1:=X41;
CylinderIO12309.xPresentDetect2:=X42;

Conveyor12114(ConveyorMotor:=ConveyorIO12114);
ConveyorIO12114.xForward:=M32;
ConveyorIO12114.xCWPresent:=X45;
Y23E:=ConveyorIO12114.xMotorCW;
M300:=NOT ConveyorIO12114.xEmpty;
M301:=ConveyorIO12114.xError;
ConveyorIO12114.iDeviceID:=12114;

Conveyor12115(ConveyorMotor:=ConveyorIO12115);
ConveyorIO12115.xForward:=M33;
ConveyorIO12115.xCWPresent:=X46;
Y23F:=ConveyorIO12115.xMotorCW;
M302:=NOT ConveyorIO12115.xEmpty;
M303:=ConveyorIO12115.xError;
ConveyorIO12115.iDeviceID:=12115;

Switch12312(ConveyorEntryIO:=ConveyorIO12116 ,
                                                        ConveyorExitIO:=ConveyorIO12123 ,
                                                        SwitchIO:=SwitchIO12312 );
SwitchIO12312.xLiftCylinderExtendButton:=M34;
SwitchIO12312.xLiftCylinderRetractButton:=M35;
Y242:=SwitchIO12312.xLiftCylinderExtend;
Y241:=SwitchIO12312.xLiftCylinderRetract;
SwitchIO12312.xLiftCylinderExtendDetect:=X4B;
SwitchIO12312.xLiftCylinderRetractDetect:=X4C;
ConveyorIO12116.xForward:=M36;
ConveyorIO12116.xCWPresent:=X49 OR X4A;
Y240:=ConveyorIO12116.xMotorCW;
M304:=NOT ConveyorIO12116.xEmpty;
M305:=ConveyorIO12116.xError;
ConveyorIO12116.iDeviceID:=12116;
ConveyorIO12123.xForward:=M37;
ConveyorIO12123.xCWPresent:=X49 OR X4A;
Y243:=ConveyorIO12123.xMotorCW;
ConveyorIO12116.tLoadDelay:=T#1s;
ConveyorIO12123.tLoadDelay:=T#2s;
M306:=NOT ConveyorIO12123.xEmpty;
M307:=ConveyorIO12123.xError;
ConveyorIO12123.iDeviceID:=12123;

Conveyor12124(ConveyorMotor:=ConveyorIO12124);
ConveyorIO12124.xForward:=M38;
ConveyorIO12124.xCWPresent:=X4D;
Y244:=conveyorIO12124.xMotorCW;
M308:=NOT ConveyorIO12124.xEmpty;
M309:=ConveyorIO12124.xError;
ConveyorIO12124.iDeviceID:=12124;

Conveyor12125(ConveyorMotor:=ConveyorIO12125);
ConveyorIO12125.xForward:=M39;
ConveyorIO12125.xCWPresent:=X4E;
Y245:=conveyorIO12125.xMotorCW;
M310:=NOT ConveyorIO12125.xEmpty;
M311:=ConveyorIO12125.xError;
ConveyorIO12125.iDeviceID:=12125;

(*常温库2巷道出库线体*)
Cylinder12308(ShuttleCarInOut:=CylinderIO12308);
ShuttleCarCurrentPosition( X35 OR X36 ,X36 ,X35, FALSE, CylinderIO12308.iCurrentPos );
CylinderIO12308.xForward:=M40;
CylinderIO12308.xBackward:=M41;
CylinderIO12308.xCylinder:=1;
Y235:=CylinderIO12308.xCW;
Y236:=CylinderIO12308.xCCW;
CylinderIO12308.xPresentDetect1:=X34;
CylinderIO12308.xPresentDetect2:=X33;

Conveyor12111(ConveyorMotor:=ConveyorIO12111);
ConveyorIO12111.xForward:=M42;
ConveyorIO12111.xCWPresent:=X37;
Y237:=ConveyorIO12111.xMotorCW;
M312:=NOT ConveyorIO12111.xEmpty;
M313:=ConveyorIO12111.xError;
ConveyorIO12111.iDeviceID:=12111;

Conveyor12112(ConveyorMotor:=ConveyorIO12112);
ConveyorIO12112.xForward:=M43;
ConveyorIO12112.xCWPresent:=X38;
Y238:=ConveyorIO12112.xMotorCW;
M314:=NOT ConveyorIO12112.xEmpty;
M315:=ConveyorIO12112.xError;
ConveyorIO12112.iDeviceID:=12112;

Switch12311(ConveyorEntryIO:=ConveyorIO12113 ,
                                                        ConveyorExitIO:=ConveyorIO12120 ,
                                                        SwitchIO:=SwitchIO12311 );
SwitchIO12311.xLiftCylinderExtendButton:=M44;
SwitchIO12311.xLiftCylinderRetractButton:=M45;
Y233:=SwitchIO12311.xLiftCylinderExtend;
Y232:=SwitchIO12311.xLiftCylinderRetract;
SwitchIO12311.xLiftCylinderExtendDetect:=X3D;
SwitchIO12311.xLiftCylinderRetractDetect:=X3E;
ConveyorIO12113.xForward:=M46;
ConveyorIO12113.xCWPresent:=X3B OR X3C;
Y239:=ConveyorIO12113.xMotorCW;
M316:=NOT ConveyorIO12113.xEmpty;
M317:=ConveyorIO12113.xError;
ConveyorIO12113.iDeviceID:=12113;
ConveyorIO12120.xForward:=M47;
ConveyorIO12120.xCWPresent:=X3B OR X3C;
Y234:=ConveyorIO12120.xMotorCW;
ConveyorIO12113.tLoadDelay:=T#1s;
ConveyorIO12120.tLoadDelay:=T#2s;
M318:=NOT ConveyorIO12120.xEmpty;
M319:=ConveyorIO12120.xError;
ConveyorIO12120.iDeviceID:=12120;

Conveyor12121(ConveyorMotor:=ConveyorIO12121);
ConveyorIO12121.xForward:=M48;
ConveyorIO12121.xCWPresent:=X3F;
Y23A:=conveyorIO12121.xMotorCW;
M320:=NOT ConveyorIO12121.xEmpty;
M321:=ConveyorIO12121.xError;
ConveyorIO12121.iDeviceID:=12121;

Conveyor12122(ConveyorMotor:=ConveyorIO12122);
ConveyorIO12122.xForward:=M49;
ConveyorIO12122.xCWPresent:=X40;
Y23B:=conveyorIO12122.xMotorCW;
M322:=NOT ConveyorIO12122.xEmpty;
M323:=ConveyorIO12122.xError;
ConveyorIO12122.iDeviceID:=12122;

(*常温库3巷道出库线体*)
Cylinder12307(ShuttleCarInOut:=CylinderIO12307);
ShuttleCarCurrentPosition( X27 OR X28 ,X28 ,X27, FALSE, CylinderIO12307.iCurrentPos );
CylinderIO12307.xForward:=M50;
CylinderIO12307.xBackward:=M51;
CylinderIO12307.xCylinder:=1;
Y229:=CylinderIO12307.xCW;
Y228:=CylinderIO12307.xCCW;
CylinderIO12307.xPresentDetect1:=X25;
CylinderIO12307.xPresentDetect2:=X26;

Conveyor12108(ConveyorMotor:=ConveyorIO12108);
ConveyorIO12108.xForward:=M52;
ConveyorIO12108.xCWPresent:=X2A;
Y22B:=ConveyorIO12108.xMotorCW;
M324:=NOT ConveyorIO12108.xEmpty;
M325:=ConveyorIO12108.xError;
ConveyorIO12108.iDeviceID:=12108;

Conveyor12109(ConveyorMotor:=ConveyorIO12109);
ConveyorIO12109.xForward:=M53;
ConveyorIO12109.xCWPresent:=X29;
Y22A:=ConveyorIO12109.xMotorCW;
M326:=NOT ConveyorIO12109.xEmpty;
M327:=ConveyorIO12109.xError;
ConveyorIO12109.iDeviceID:=12109;